// TIA Portal project "Hydroelectric Power Plant" (V20) (continued)
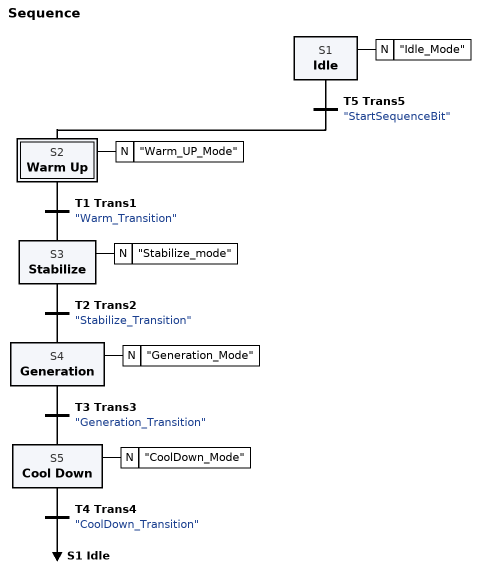
   // sequencer 1
   INITIAL_STEP "Warm Up":   // S2, max time T#10S, warning time T#7S
              N    "Warm_UP_Mode"
   END_STEP
   TRANSITION Trans1 FROM "Warm Up" TO Stabilize   // T1
      := "Warm_Transition";
   END_TRANSITION
   STEP Stabilize:   // S3, max time T#10S, warning time T#7S
              N    "Stabilize_mode"
   END_STEP
   TRANSITION Trans2 FROM Stabilize TO Generation   // T2
      := "Stabilize_Transition";
   END_TRANSITION
   STEP Generation:   // S4, max time T#10S, warning time T#7S
              N    "Generation_Mode"
   END_STEP
   TRANSITION Trans3 FROM Generation TO "Cool Down"   // T3
      := "Generation_Transition";
   END_TRANSITION
   STEP "Cool Down":   // S5, max time T#10S, warning time T#7S
              N    "CoolDown_Mode"
   END_STEP
   TRANSITION Trans4 FROM "Cool Down" TO Idle   // T4, jump
      := "CoolDown_Transition";
   END_TRANSITION
   STEP Idle:   // S1, max time T#10S, warning time T#7S
              N    "Idle_Mode"
   END_STEP
   TRANSITION Trans5 FROM Idle TO "Warm Up"   // T5
      := "StartSequenceBit";
   END_TRANSITION
END_FUNCTION_BLOCK

FUNCTION "Scale_with_parameter" : Void   // FC1, FBD
{ S7_Optimized_Access := 'TRUE' }
VERSION : 0.1
   VAR_INPUT
      input_min : Int;
      input_signal : Int;
      input_max : Int;
      output_max : Int;
      output_min : Int;
   END_VAR
   VAR_OUTPUT
      scaled_value : Int;
   END_VAR
   VAR_TEMP
      temp_value : Real;
   END_VAR
BEGIN

REGION Network 1
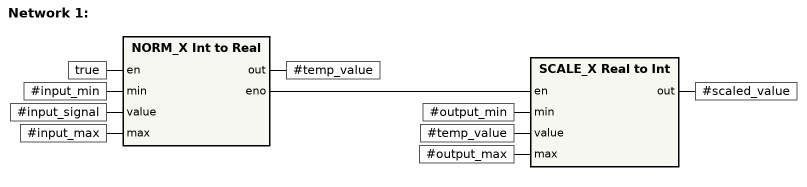
   IF true THEN
       #temp_value := NORM_X(MIN := #input_min, VALUE := #input_signal, MAX := #input_max);
       #scaled_value := SCALE_X(MIN := #output_min, VALUE := #temp_value, MAX := #output_max);
   END_IF;
END_REGION
END_FUNCTION

FUNCTION "Convert_time" : Void   // FC2, FBD
{ S7_Optimized_Access := 'TRUE' }
VERSION : 0.1
   VAR_INPUT
      iv1 : Int;
   END_VAR
   VAR_OUTPUT
      time1 : Time;
   END_VAR
   VAR_TEMP
      Int1 : Int;
   END_VAR
BEGIN

REGION Network 1
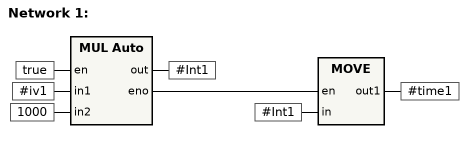
   IF true THEN
       #Int1 := #iv1 * 1000;
       #time1 := #Int1;
   END_IF;
END_REGION
END_FUNCTION

ORGANIZATION_BLOCK "Main"   // OB1, LAD, ProgramCycle
TITLE = "Main Program Sweep (Cycle)"
{ S7_Optimized_Access := 'TRUE' }
VERSION : 0.1
   VAR_INPUT
      Initial_Call : Bool;   // Initial call of this OB
      Remanence : Bool;   // =True, if remanent data are available
   END_VAR
   VAR_TEMP
      SequenceInit : Bool;
      InitSequence : Bool;
      IntSequence : Bool;
   END_VAR
   VAR_TEMP   // added for the SCL form of the ladder/FBD networks
      _w1 : Bool;
      _w2 : Bool;
      _w3 : Bool;
      _w4 : Bool;
   END_VAR
BEGIN

REGION Network 1
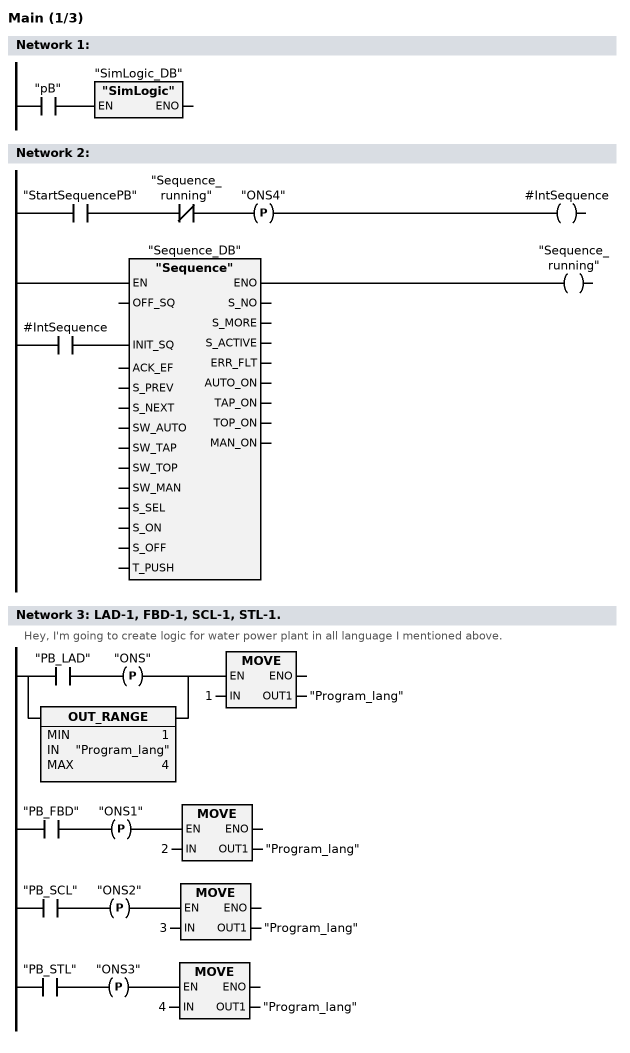
   RUNG wire#powerrail
      Contact( "pB" )
      "SimLogic_DB"()
   END_RUNG
   // the same network as SCL:
   IF "pB" THEN
       "SimLogic_DB"();   // "SimLogic"
   END_IF;
END_REGION

REGION Network 2
   RUNG wire#powerrail
      Contact( "StartSequencePB" )
      I_Contact( "Sequence_running" )
      P_Trig( "ONS4" )
      Coil( #IntSequence )
   END_RUNG
   RUNG wire#powerrail
      "Sequence_DB"(INIT_SQ := wire#w1, OFF_SQ :=, ACK_EF :=, S_PREV :=, S_NEXT :=, SW_AUTO :=, SW_TAP :=, SW_TOP :=, SW_MAN :=, S_SEL :=, S_ON :=, S_OFF :=, T_PUSH :=, S_NO =>, S_MORE =>, S_ACTIVE =>, ERR_FLT =>, AUTO_ON =>, TAP_ON =>, TOP_ON =>, MAN_ON =>)
      Coil( "Sequence_running" )
   END_RUNG
   RUNG wire#powerrail
      Contact( #IntSequence )
   END_RUNG wire#w1
   // the same network as SCL:
   #_w1 := "StartSequencePB" AND NOT "Sequence_running";
   #_w2 := #_w1 AND NOT "ONS4";   // rising edge
   "ONS4" := #_w1;
   #IntSequence := #_w2;
   "Sequence_DB"(INIT_SQ := #IntSequence, ENO => #_w3);   // "Sequence"
   "Sequence_running" := #_w3;
END_REGION

REGION Network 3: LAD-1, FBD-1, SCL-1, STL-1.
   // Hey, I'm going to create logic for water power plant in all language I mentioned above.
   #_w1 := "PB_LAD" AND NOT "ONS";   // rising edge
   "ONS" := "PB_LAD";
   IF #_w1 OR ("Program_lang" < 1) OR ("Program_lang" > 4) THEN "Program_lang" := 1; END_IF;
   #_w2 := "PB_FBD" AND NOT "ONS1";   // rising edge
   "ONS1" := "PB_FBD";
   IF #_w2 THEN "Program_lang" := 2; END_IF;
   #_w3 := "PB_SCL" AND NOT "ONS2";   // rising edge
   "ONS2" := "PB_SCL";
   IF #_w3 THEN "Program_lang" := 3; END_IF;
   #_w4 := "PB_STL" AND NOT "ONS3";   // rising edge
   "ONS3" := "PB_STL";
   IF #_w4 THEN "Program_lang" := 4; END_IF;
END_REGION

REGION Network 4: I/O for LAD
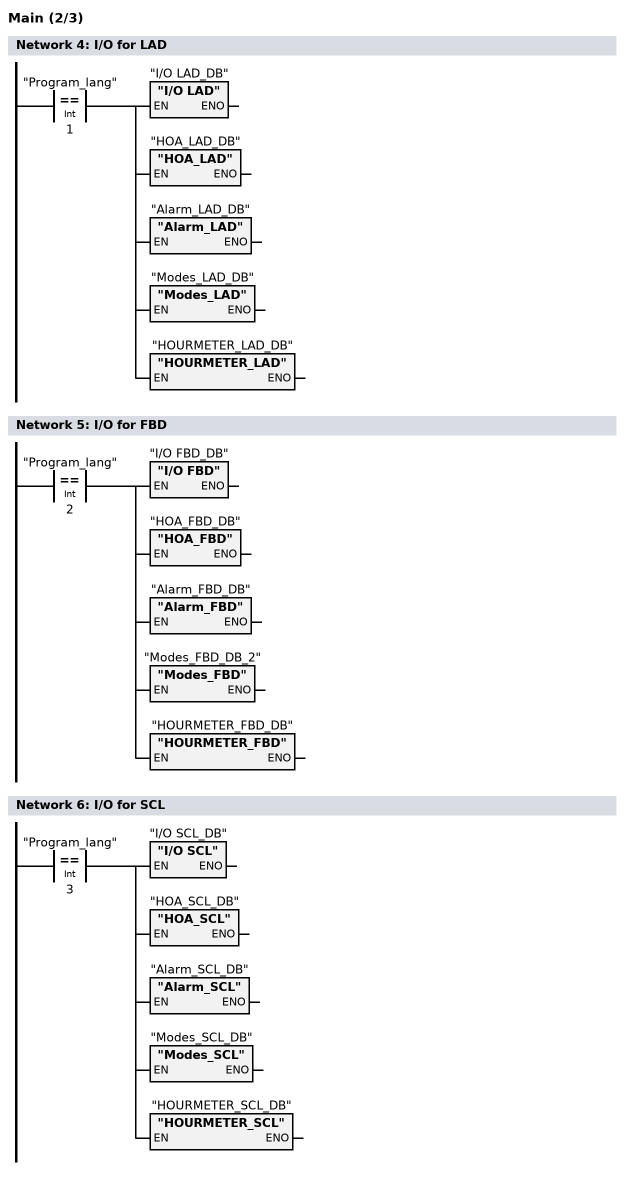
   RUNG wire#powerrail
      { S7_Templates := "SrcType := Int" } EQ_Contact(in1 := "Program_lang", in2 := 1)
      wire#w1
      "I/O LAD_DB"()
   END_RUNG
   RUNG wire#w1
      "HOA_LAD_DB"()
   END_RUNG
   RUNG wire#w1
      "Alarm_LAD_DB"()
   END_RUNG
   RUNG wire#w1
      "Modes_LAD_DB"()
   END_RUNG
   RUNG wire#w1
      "HOURMETER_LAD_DB"()
   END_RUNG
   // the same network as SCL:
   #_w1 := "Program_lang" = 1;
   IF #_w1 THEN
       "I/O LAD_DB"();   // "I/O LAD"
       "HOA_LAD_DB"();   // "HOA_LAD"
       "Alarm_LAD_DB"();   // "Alarm_LAD"
       "Modes_LAD_DB"();   // "Modes_LAD"
       "HOURMETER_LAD_DB"();   // "HOURMETER_LAD"
   END_IF;
END_REGION

REGION Network 5: I/O for FBD
   RUNG wire#powerrail
      { S7_Templates := "SrcType := Int" } EQ_Contact(in1 := "Program_lang", in2 := 2)
      wire#w1
      "I/O FBD_DB"()
   END_RUNG
   RUNG wire#w1
      "HOA_FBD_DB"()
   END_RUNG
   RUNG wire#w1
      "Alarm_FBD_DB"()
   END_RUNG
   RUNG wire#w1
      "Modes_FBD_DB_2"()
   END_RUNG
   RUNG wire#w1
      "HOURMETER_FBD_DB"()
   END_RUNG
   // the same network as SCL:
   #_w1 := "Program_lang" = 2;
   IF #_w1 THEN
       "I/O FBD_DB"();   // "I/O FBD"
       "HOA_FBD_DB"();   // "HOA_FBD"
       "Alarm_FBD_DB"();   // "Alarm_FBD"
       "Modes_FBD_DB_2"();   // "Modes_FBD"
       "HOURMETER_FBD_DB"();   // "HOURMETER_FBD"
   END_IF;
END_REGION

REGION Network 6: I/O for SCL
   RUNG wire#powerrail
      { S7_Templates := "SrcType := Int" } EQ_Contact(in1 := "Program_lang", in2 := 3)
      wire#w1
      "I/O SCL_DB"()
   END_RUNG
   RUNG wire#w1
      "HOA_SCL_DB"()
   END_RUNG
   RUNG wire#w1
      "Alarm_SCL_DB"()
   END_RUNG
   RUNG wire#w1
      "Modes_SCL_DB"()
   END_RUNG
   RUNG wire#w1
      "HOURMETER_SCL_DB"()
   END_RUNG
   // the same network as SCL:
   #_w1 := "Program_lang" = 3;
   IF #_w1 THEN
       "I/O SCL_DB"();   // "I/O SCL"
       "HOA_SCL_DB"();   // "HOA_SCL"
       "Alarm_SCL_DB"();   // "Alarm_SCL"
       "Modes_SCL_DB"();   // "Modes_SCL"
       "HOURMETER_SCL_DB"();   // "HOURMETER_SCL"
   END_IF;
END_REGION

REGION Network 7: I/O for STL
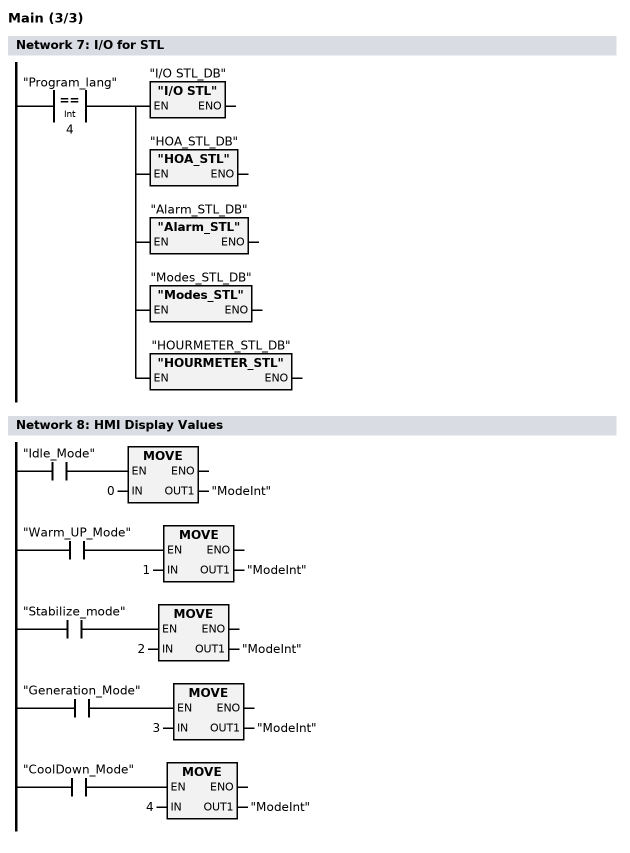
   RUNG wire#powerrail
      { S7_Templates := "SrcType := Int" } EQ_Contact(in1 := "Program_lang", in2 := 4)
      wire#w1
      "I/O STL_DB"()
   END_RUNG
   RUNG wire#w1
      "HOA_STL_DB"()
   END_RUNG
   RUNG wire#w1
      "Alarm_STL_DB"()
   END_RUNG
   RUNG wire#w1
      "Modes_STL_DB"()
   END_RUNG
   RUNG wire#w1
      "HOURMETER_STL_DB"()
   END_RUNG
   // the same network as SCL:
   #_w1 := "Program_lang" = 4;
   IF #_w1 THEN
       "I/O STL_DB"();   // "I/O STL"
       "HOA_STL_DB"();   // "HOA_STL"
       "Alarm_STL_DB"();   // "Alarm_STL"
       "Modes_STL_DB"();   // "Modes_STL"
       "HOURMETER_STL_DB"();   // "HOURMETER_STL"
   END_IF;
END_REGION

REGION Network 8: HMI Display Values
   RUNG wire#powerrail
      Contact( "Idle_Mode" )
      Move(in := 0, out1 => "ModeInt")
   END_RUNG
   RUNG wire#powerrail
      Contact( "Warm_UP_Mode" )
      Move(in := 1, out1 => "ModeInt")
   END_RUNG
   RUNG wire#powerrail
      Contact( "Stabilize_mode" )
      Move(in := 2, out1 => "ModeInt")
   END_RUNG
   RUNG wire#powerrail
      Contact( "Generation_Mode" )
      Move(in := 3, out1 => "ModeInt")
   END_RUNG
   RUNG wire#powerrail
      Contact( "CoolDown_Mode" )
      Move(in := 4, out1 => "ModeInt")
   END_RUNG
   // the same network as SCL:
   IF "Idle_Mode" THEN "ModeInt" := 0; END_IF;
   IF "Warm_UP_Mode" THEN "ModeInt" := 1; END_IF;
   IF "Stabilize_mode" THEN "ModeInt" := 2; END_IF;
   IF "Generation_Mode" THEN "ModeInt" := 3; END_IF;
   IF "CoolDown_Mode" THEN "ModeInt" := 4; END_IF;
END_REGION
END_ORGANIZATION_BLOCK

ORGANIZATION_BLOCK "PID"   // OB30, LAD, CyclicInterrupt
{ S7_Optimized_Access := 'TRUE' }
VERSION : 0.1
   VAR_INPUT
      Initial_Call : Bool;   // Initial call of this OB
      Event_Count : Int;   // Events discarded
   END_VAR
   VAR_TEMP
      Bsp : Real;
      Vsp : Real;
      bafflehand_trigger : Bool;
      baffleoff_trigger : Bool;
      baffleauto_trigger : Bool;
      vfdhand_trigger : Bool;
      vfdoff_trigger : Bool;
      vfdauto_trigger : Bool;
   END_VAR
   VAR_TEMP   // added for the SCL form of the ladder/FBD networks
      _w1 : Bool;
      _w2 : Bool;
      _w3 : Bool;
      _w4 : Bool;
      _w5 : Bool;
      _w6 : Bool;
      _w7 : Bool;
   END_VAR
BEGIN

REGION Network 1: high oil flow alarm handling
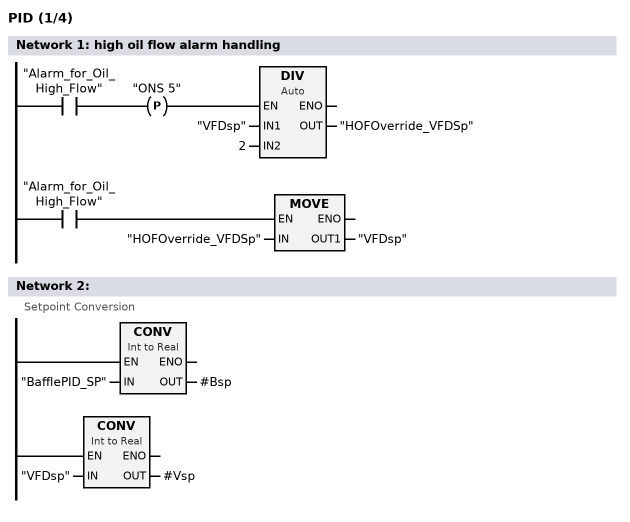
   RUNG wire#powerrail
      Contact( "Alarm_for_Oil_High_Flow" )
      P_Trig( "ONS 5" )
      Div(in1 := "VFDsp", in2 := 2, out => "HOFOverride_VFDSp")
   END_RUNG
   RUNG wire#powerrail
      Contact( "Alarm_for_Oil_High_Flow" )
      Move(in := "HOFOverride_VFDSp", out1 => "VFDsp")
   END_RUNG
   // the same network as SCL:
   #_w1 := "Alarm_for_Oil_High_Flow" AND NOT "ONS 5";   // rising edge
   "ONS 5" := "Alarm_for_Oil_High_Flow";
   IF #_w1 THEN "HOFOverride_VFDSp" := "VFDsp" / 2; END_IF;
   IF "Alarm_for_Oil_High_Flow" THEN "VFDsp" := "HOFOverride_VFDSp"; END_IF;
END_REGION

REGION Network 2
   // Setpoint Conversion
   RUNG wire#powerrail
      { S7_Templates := "[SrcType := Int, DestType := Real]" } Convert(in := "BafflePID_SP", out => #Bsp)
   END_RUNG
   RUNG wire#powerrail
      { S7_Templates := "[SrcType := Int, DestType := Real]" } Convert(in := "VFDsp", out => #Vsp)
   END_RUNG
   // the same network as SCL:
   #Bsp := INT_TO_REAL("BafflePID_SP");
   #Vsp := INT_TO_REAL("VFDsp");
END_REGION

REGION Network 3
   // Baffle HOA
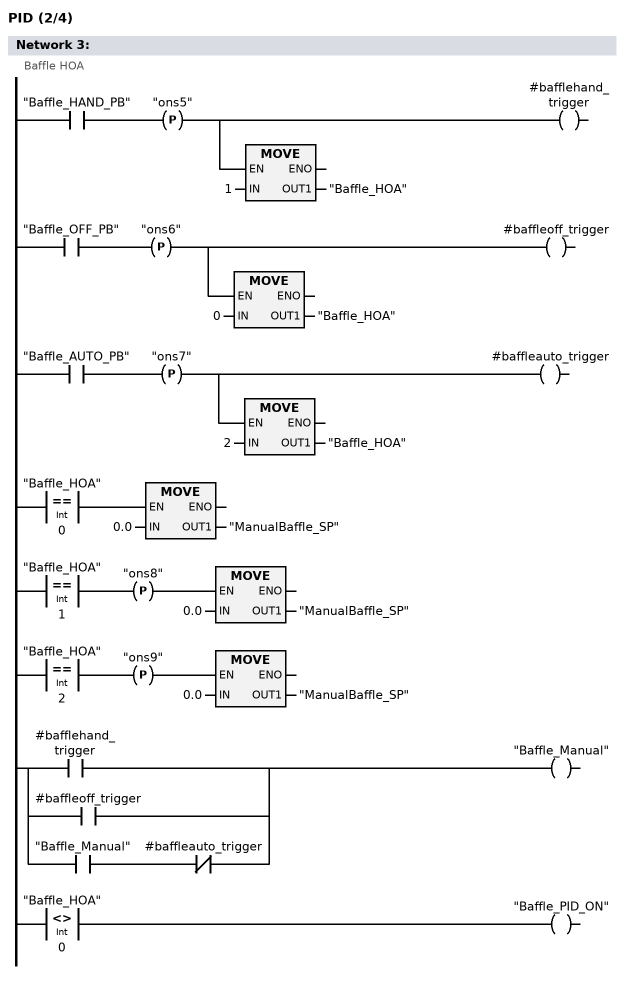
   RUNG wire#powerrail
      Contact( "Baffle_HAND_PB" )
      P_Trig( "ons5" )
      wire#w1
      Coil( #bafflehand_trigger )
   END_RUNG
   RUNG wire#w1
      Move(in := 1, out1 => "Baffle_HOA")
   END_RUNG
   RUNG wire#powerrail
      Contact( "Baffle_OFF_PB" )
      P_Trig( "ons6" )
      wire#w2
      Coil( #baffleoff_trigger )
   END_RUNG
   RUNG wire#w2
      Move(in := 0, out1 => "Baffle_HOA")
   END_RUNG
   RUNG wire#powerrail
      Contact( "Baffle_AUTO_PB" )
      P_Trig( "ons7" )
      wire#w3
      Coil( #baffleauto_trigger )
   END_RUNG
   RUNG wire#w3
      Move(in := 2, out1 => "Baffle_HOA")
   END_RUNG
   RUNG wire#powerrail
      { S7_Templates := "SrcType := Int" } EQ_Contact(in1 := "Baffle_HOA", in2 := 0)
      Move(in := 0.0, out1 => "ManualBaffle_SP")
   END_RUNG
   RUNG wire#powerrail
      { S7_Templates := "SrcType := Int" } EQ_Contact(in1 := "Baffle_HOA", in2 := 1)
      P_Trig( "ons8" )
      Move(in := 0.0, out1 => "ManualBaffle_SP")
   END_RUNG
   RUNG wire#powerrail
      { S7_Templates := "SrcType := Int" } EQ_Contact(in1 := "Baffle_HOA", in2 := 2)
      P_Trig( "ons9" )
      Move(in := 0.0, out1 => "ManualBaffle_SP")
   END_RUNG
   RUNG wire#powerrail
      Contact( #bafflehand_trigger )
      wire#w4
      Coil( "Baffle_Manual" )
   END_RUNG
   RUNG wire#powerrail
      Contact( #baffleoff_trigger )
   END_RUNG wire#w4
   RUNG wire#powerrail
      Contact( "Baffle_Manual" )
      I_Contact( #baffleauto_trigger )
   END_RUNG wire#w4
   RUNG wire#powerrail
      { S7_Templates := "SrcType := Int" } NE_Contact(in1 := "Baffle_HOA", in2 := 0)
      Coil( "Baffle_PID_ON" )
   END_RUNG
   // the same network as SCL:
   #_w1 := "Baffle_HAND_PB" AND NOT "ons5";   // rising edge
   "ons5" := "Baffle_HAND_PB";
   #bafflehand_trigger := #_w1;
   IF #_w1 THEN "Baffle_HOA" := 1; END_IF;
   #_w2 := "Baffle_OFF_PB" AND NOT "ons6";   // rising edge
   "ons6" := "Baffle_OFF_PB";
   #baffleoff_trigger := #_w2;
   IF #_w2 THEN "Baffle_HOA" := 0; END_IF;
   #_w3 := "Baffle_AUTO_PB" AND NOT "ons7";   // rising edge
   "ons7" := "Baffle_AUTO_PB";
   #baffleauto_trigger := #_w3;
   IF #_w3 THEN "Baffle_HOA" := 2; END_IF;
   IF "Baffle_HOA" = 0 THEN "ManualBaffle_SP" := 0.0; END_IF;
   #_w4 := "Baffle_HOA" = 1;
   #_w5 := #_w4 AND NOT "ons8";   // rising edge
   "ons8" := #_w4;
   IF #_w5 THEN "ManualBaffle_SP" := 0.0; END_IF;
   #_w6 := "Baffle_HOA" = 2;
   #_w7 := #_w6 AND NOT "ons9";   // rising edge
   "ons9" := #_w6;
   IF #_w7 THEN "ManualBaffle_SP" := 0.0; END_IF;
   "Baffle_Manual" := #bafflehand_trigger OR #baffleoff_trigger OR ("Baffle_Manual" AND NOT #baffleauto_trigger);
   "Baffle_PID_ON" := "Baffle_HOA" <> 0;
END_REGION

REGION Network 4
   // VFD HOA
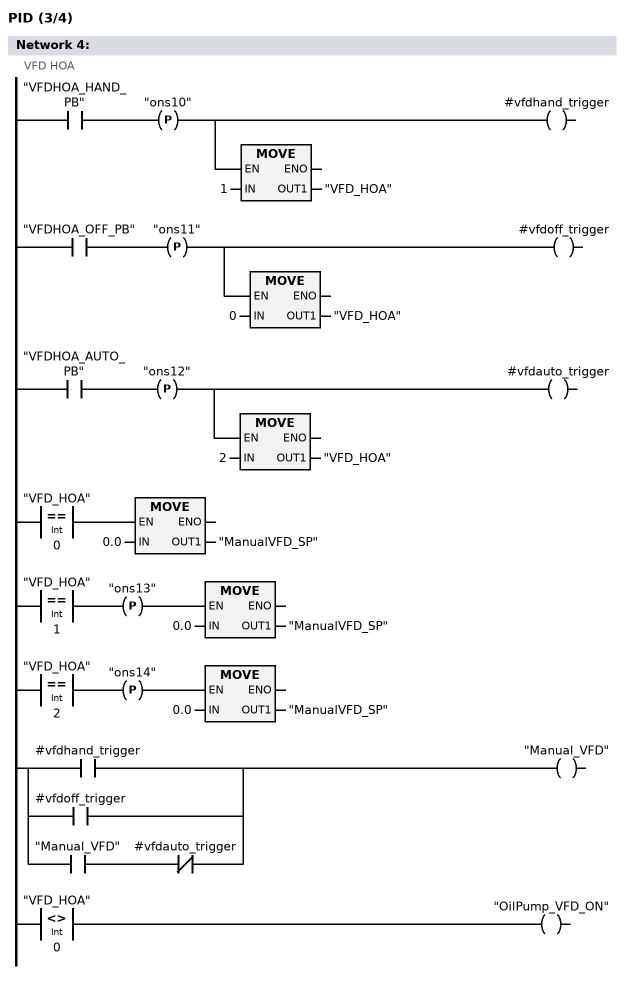
   RUNG wire#powerrail
      Contact( "VFDHOA_HAND_PB" )
      P_Trig( "ons10" )
      wire#w1
      Coil( #vfdhand_trigger )
   END_RUNG
   RUNG wire#w1
      Move(in := 1, out1 => "VFD_HOA")
   END_RUNG
   RUNG wire#powerrail
      Contact( "VFDHOA_OFF_PB" )
      P_Trig( "ons11" )
      wire#w2
      Coil( #vfdoff_trigger )
   END_RUNG
   RUNG wire#w2
      Move(in := 0, out1 => "VFD_HOA")
   END_RUNG
   RUNG wire#powerrail
      Contact( "VFDHOA_AUTO_PB" )
      P_Trig( "ons12" )
      wire#w3
      Coil( #vfdauto_trigger )
   END_RUNG
   RUNG wire#w3
      Move(in := 2, out1 => "VFD_HOA")
   END_RUNG
   RUNG wire#powerrail
      { S7_Templates := "SrcType := Int" } EQ_Contact(in1 := "VFD_HOA", in2 := 0)
      Move(in := 0.0, out1 => "ManualVFD_SP")
   END_RUNG
   RUNG wire#powerrail
      { S7_Templates := "SrcType := Int" } EQ_Contact(in1 := "VFD_HOA", in2 := 1)
      P_Trig( "ons13" )
      Move(in := 0.0, out1 => "ManualVFD_SP")
   END_RUNG
   RUNG wire#powerrail
      { S7_Templates := "SrcType := Int" } EQ_Contact(in1 := "VFD_HOA", in2 := 2)
      P_Trig( "ons14" )
      Move(in := 0.0, out1 => "ManualVFD_SP")
   END_RUNG
   RUNG wire#powerrail
      Contact( #vfdhand_trigger )
      wire#w4
      Coil( "Manual_VFD" )
   END_RUNG
   RUNG wire#powerrail
      Contact( #vfdoff_trigger )
   END_RUNG wire#w4
   RUNG wire#powerrail
      Contact( "Manual_VFD" )
      I_Contact( #vfdauto_trigger )
   END_RUNG wire#w4
   RUNG wire#powerrail
      { S7_Templates := "SrcType := Int" } NE_Contact(in1 := "VFD_HOA", in2 := 0)
      Coil( "OilPump_VFD_ON" )
   END_RUNG
   // the same network as SCL:
   #_w1 := "VFDHOA_HAND_PB" AND NOT "ons10";   // rising edge
   "ons10" := "VFDHOA_HAND_PB";
   #vfdhand_trigger := #_w1;
   IF #_w1 THEN "VFD_HOA" := 1; END_IF;
   #_w2 := "VFDHOA_OFF_PB" AND NOT "ons11";   // rising edge
   "ons11" := "VFDHOA_OFF_PB";
   #vfdoff_trigger := #_w2;
   IF #_w2 THEN "VFD_HOA" := 0; END_IF;
   #_w3 := "VFDHOA_AUTO_PB" AND NOT "ons12";   // rising edge
   "ons12" := "VFDHOA_AUTO_PB";
   #vfdauto_trigger := #_w3;
   IF #_w3 THEN "VFD_HOA" := 2; END_IF;
   IF "VFD_HOA" = 0 THEN "ManualVFD_SP" := 0.0; END_IF;
   #_w4 := "VFD_HOA" = 1;
   #_w5 := #_w4 AND NOT "ons13";   // rising edge
   "ons13" := #_w4;
   IF #_w5 THEN "ManualVFD_SP" := 0.0; END_IF;
   #_w6 := "VFD_HOA" = 2;
   #_w7 := #_w6 AND NOT "ons14";   // rising edge
   "ons14" := #_w6;
   IF #_w7 THEN "ManualVFD_SP" := 0.0; END_IF;
   "Manual_VFD" := #vfdhand_trigger OR #vfdoff_trigger OR ("Manual_VFD" AND NOT #vfdauto_trigger);
   "OilPump_VFD_ON" := "VFD_HOA" <> 0;
END_REGION

REGION Network 5
   // PID
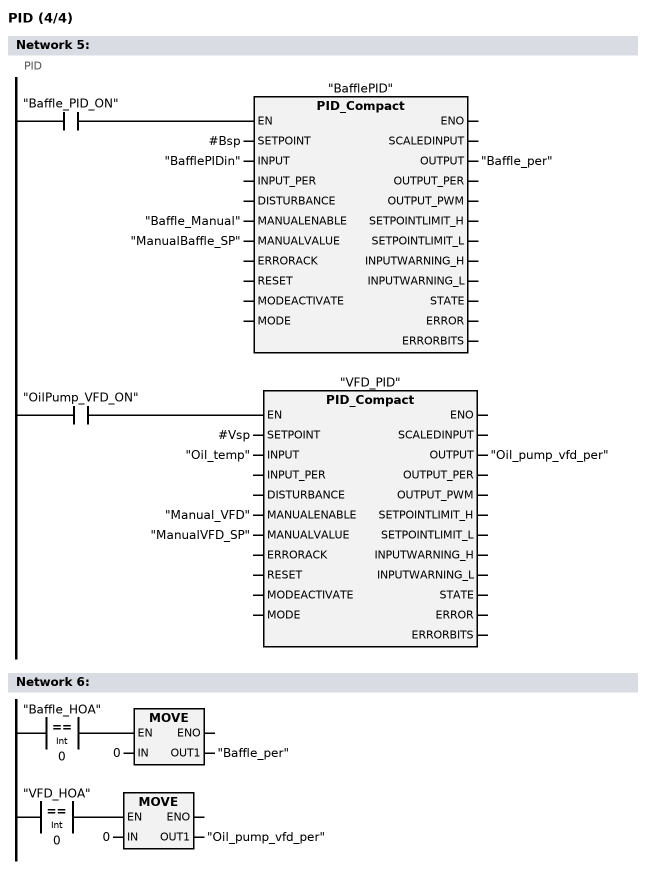
   IF "Baffle_PID_ON" THEN
       "BafflePID"(Setpoint := #Bsp,   // PID_Compact
                   Input := "BafflePIDin",
                   ManualEnable := "Baffle_Manual",
                   ManualValue := "ManualBaffle_SP",
                   Output => "Baffle_per");
   END_IF;
   IF "OilPump_VFD_ON" THEN
       "VFD_PID"(Setpoint := #Vsp,   // PID_Compact
                 Input := "Oil_temp",
                 ManualEnable := "Manual_VFD",
                 ManualValue := "ManualVFD_SP",
                 Output => "Oil_pump_vfd_per");
   END_IF;
END_REGION

REGION Network 6
   RUNG wire#powerrail
      { S7_Templates := "SrcType := Int" } EQ_Contact(in1 := "Baffle_HOA", in2 := 0)
      Move(in := 0, out1 => "Baffle_per")
   END_RUNG
   RUNG wire#powerrail
      { S7_Templates := "SrcType := Int" } EQ_Contact(in1 := "VFD_HOA", in2 := 0)
      Move(in := 0, out1 => "Oil_pump_vfd_per")
   END_RUNG
   // the same network as SCL:
   IF "Baffle_HOA" = 0 THEN "Baffle_per" := 0; END_IF;
   IF "VFD_HOA" = 0 THEN "Oil_pump_vfd_per" := 0; END_IF;
END_REGION
END_ORGANIZATION_BLOCK

// folder: FBD

FUNCTION_BLOCK "I/O FBD"   // FB3, FBD
TITLE = FBD I/O and Scaling parameters
{ S7_Optimized_Access := 'TRUE' }
VERSION : 0.1
   VAR_TEMP
      Temp_v : Real;
   END_VAR
BEGIN

REGION Network 1: Digital Output's
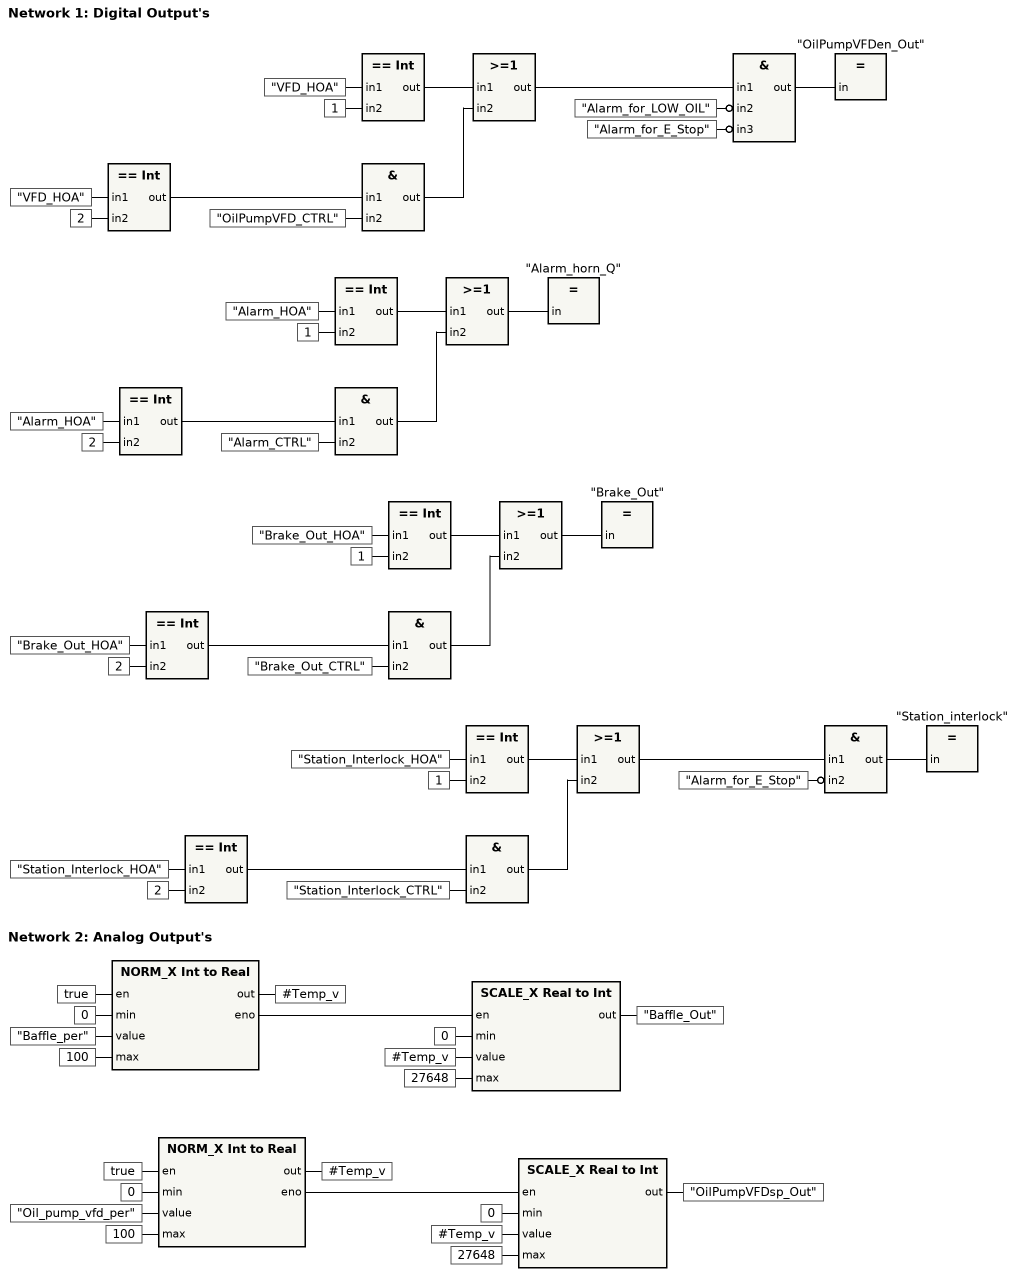
   "OilPumpVFDen_Out" := (("VFD_HOA" = 1) OR (("VFD_HOA" = 2) AND "OilPumpVFD_CTRL")) AND NOT "Alarm_for_LOW_OIL" AND NOT "Alarm_for_E_Stop";
   "Alarm_horn_Q" := ("Alarm_HOA" = 1) OR (("Alarm_HOA" = 2) AND "Alarm_CTRL");
   "Brake_Out" := ("Brake_Out_HOA" = 1) OR (("Brake_Out_HOA" = 2) AND "Brake_Out_CTRL");
   "Station_interlock" := (("Station_Interlock_HOA" = 1) OR (("Station_Interlock_HOA" = 2) AND "Station_Interlock_CTRL")) AND NOT "Alarm_for_E_Stop";
END_REGION

REGION Network 2: Analog Output's
   IF true THEN
       #Temp_v := NORM_X(MIN := 0, VALUE := "Baffle_per", MAX := 100);
       "Baffle_Out" := SCALE_X(MIN := 0, VALUE := #Temp_v, MAX := 27648);
       #Temp_v := NORM_X(MIN := 0, VALUE := "Oil_pump_vfd_per", MAX := 100);
       "OilPumpVFDsp_Out" := SCALE_X(MIN := 0, VALUE := #Temp_v, MAX := 27648);
   END_IF;
END_REGION

REGION Network 3: Analog Input's
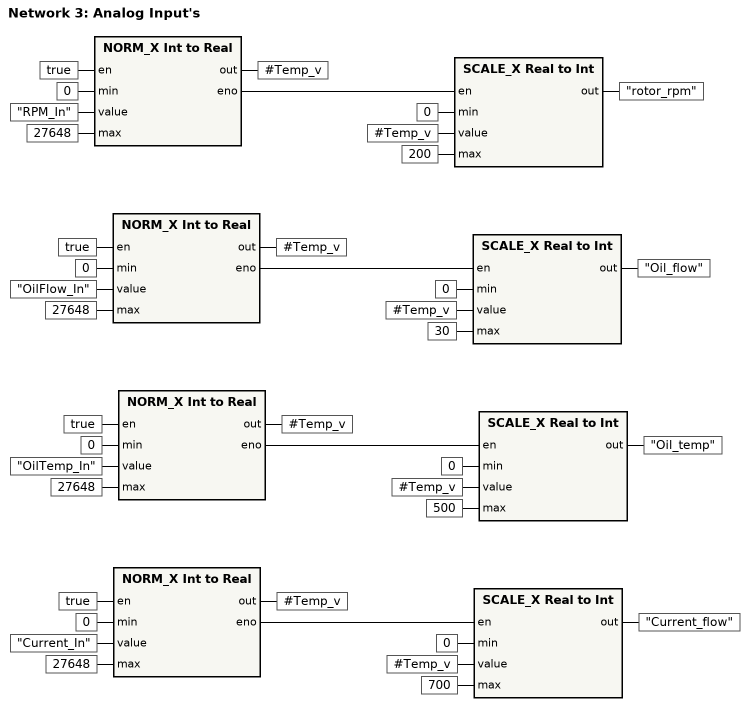
   IF true THEN
       #Temp_v := NORM_X(MIN := 0, VALUE := "RPM_In", MAX := 27648);
       "rotor_rpm" := SCALE_X(MIN := 0, VALUE := #Temp_v, MAX := 200);
       #Temp_v := NORM_X(MIN := 0, VALUE := "OilFlow_In", MAX := 27648);
       "Oil_flow" := SCALE_X(MIN := 0, VALUE := #Temp_v, MAX := 30);
       #Temp_v := NORM_X(MIN := 0, VALUE := "OilTemp_In", MAX := 27648);
       "Oil_temp" := SCALE_X(MIN := 0, VALUE := #Temp_v, MAX := 500);
       #Temp_v := NORM_X(MIN := 0, VALUE := "Current_In", MAX := 27648);
       "Current_flow" := SCALE_X(MIN := 0, VALUE := #Temp_v, MAX := 700);
   END_IF;
END_REGION

REGION Network 4
   // FULLAUTOBIT
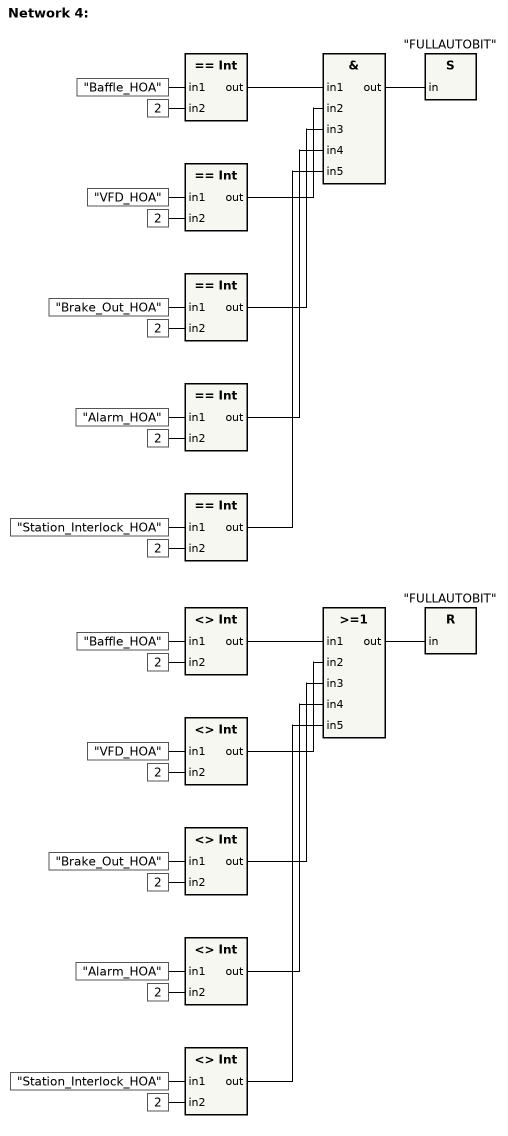
   IF ("Baffle_HOA" = 2) AND ("VFD_HOA" = 2) AND ("Brake_Out_HOA" = 2) AND ("Alarm_HOA" = 2) AND ("Station_Interlock_HOA" = 2) THEN
       "FULLAUTOBIT" := TRUE;
   END_IF;
   IF ("Baffle_HOA" <> 2) OR ("VFD_HOA" <> 2) OR ("Brake_Out_HOA" <> 2) OR ("Alarm_HOA" <> 2) OR ("Station_Interlock_HOA" <> 2) THEN
       "FULLAUTOBIT" := FALSE;
   END_IF;
END_REGION
END_FUNCTION_BLOCK

FUNCTION_BLOCK "HOA_FBD"   // FB7, FBD
{ S7_Optimized_Access := 'TRUE' }